   Button "Schaltfläche_256" at 1154,453 size 59x15; TextOff 'Text'
      on Click: SetTag("_DB_SDC_ERRORS.Error_nr", 830)
   Button "Schaltfläche_257" at 1154,469 size 59x15; TextOff 'Text'
      on Click: SetTag("_DB_SDC_ERRORS.Error_nr", 831)
   Button "Schaltfläche_258" at 1154,485 size 59x15; TextOff 'Text'
      on Click: SetTag("_DB_SDC_ERRORS.Error_nr", 832)
   Button "Schaltfläche_259" at 971,533 size 59x15; TextOff 'Text'
      on Click: SetTag("_DB_SDC_ERRORS.Error_nr", 901)
   Button "Schaltfläche_260" at 971,549 size 59x15; TextOff 'Text'
      on Click: SetTag("_DB_SDC_ERRORS.Error_nr", 902)
   Button "Schaltfläche_261" at 971,565 size 59x15; TextOff 'Text'
      on Click: SetTag("_DB_SDC_ERRORS.Error_nr", 903)
   Button "Schaltfläche_262" at 971,581 size 59x15; TextOff 'Text'
      on Click: SetTag("_DB_SDC_ERRORS.Error_nr", 904)
   Button "Schaltfläche_263" at 971,597 size 59x15; TextOff 'Text'
      on Click: SetTag("_DB_SDC_ERRORS.Error_nr", 905)
   Button "Schaltfläche_264" at 971,613 size 59x15; TextOff 'Text'
      on Click: SetTag("_DB_SDC_ERRORS.Error_nr", 906)
   Button "Schaltfläche_265" at 971,629 size 59x15; TextOff 'Text'
      on Click: SetTag("_DB_SDC_ERRORS.Error_nr", 907)
   Button "Schaltfläche_266" at 971,645 size 59x15; TextOff 'Text'
      on Click: SetTag("_DB_SDC_ERRORS.Error_nr", 908)
   Button "Schaltfläche_267" at 1033,533 size 59x15; TextOff 'Text'
      on Click: SetTag("_DB_SDC_ERRORS.Error_nr", 909)
   Button "Schaltfläche_268" at 1033,549 size 59x15; TextOff 'Text'
      on Click: SetTag("_DB_SDC_ERRORS.Error_nr", 910)
   Button "Schaltfläche_269" at 1033,565 size 59x15; TextOff 'Text'
      on Click: SetTag("_DB_SDC_ERRORS.Error_nr", 911)
   Button "Schaltfläche_270" at 1033,581 size 59x15; TextOff 'Text'
      on Click: SetTag("_DB_SDC_ERRORS.Error_nr", 912)
   Button "Schaltfläche_271" at 1033,597 size 59x15; TextOff 'Text'
      on Click: SetTag("_DB_SDC_ERRORS.Error_nr", 913)
   Button "Schaltfläche_272" at 1033,613 size 59x15; TextOff 'Text'
      on Click: SetTag("_DB_SDC_ERRORS.Error_nr", 914)
   Button "Schaltfläche_273" at 1033,629 size 59x15; TextOff 'Text'
      on Click: SetTag("_DB_SDC_ERRORS.Error_nr", 915)
   Button "Schaltfläche_274" at 1033,645 size 59x15; TextOff 'Text'
      on Click: SetTag("_DB_SDC_ERRORS.Error_nr", 916)
   Button "Schaltfläche_275" at 977,670 size 54x15; TextOff 'Text'
      on Click: SetTag("_DB_SDC_ERRORS.Error_nr", 917)
   Button "Schaltfläche_276" at 977,686 size 54x15; TextOff 'Text'
      on Click: SetTag("_DB_SDC_ERRORS.Error_nr", 918)
   Button "Schaltfläche_277" at 977,702 size 54x15; TextOff 'Text'
      on Click: SetTag("_DB_SDC_ERRORS.Error_nr", 919)
   Button "Schaltfläche_278" at 977,718 size 54x15; TextOff 'Text'
      on Click: SetTag("_DB_SDC_ERRORS.Error_nr", 920)
   Button "Schaltfläche_279" at 1032,669 size 54x15; TextOff 'Text'
      on Click: SetTag("_DB_SDC_ERRORS.Error_nr", 921)
   Button "Schaltfläche_280" at 1032,685 size 54x15; TextOff 'Text'
      on Click: SetTag("_DB_SDC_ERRORS.Error_nr", 922)
   Button "Schaltfläche_281" at 1032,701 size 54x15; TextOff 'Text'
      on Click: SetTag("_DB_SDC_ERRORS.Error_nr", 923)
   Button "Schaltfläche_282" at 1032,717 size 54x15; TextOff 'Text'
      on Click: SetTag("_DB_SDC_ERRORS.Error_nr", 924)

screen "724_ERROR_STAT_NOT_USED" 1280x800, template "Top_Header"
   on GenerateScreen: "SDC_ERROR_STAT"("SDC\DB_SDC_ERROR_STAT\_intern_Fault_Stat_Nr"); SetTag("SDC\_intern_Bildnummer", 724)
   IOField "EA-Feld_1" at 372,374 size 96x27; FormatPattern 999999999
      ProcessValue <- "SDC\DB_SDC_ERROR_STAT\DB_SDC_ERROR_STAT.F_STAT[XX1].EMS_TS_STAT_VAL.DRIVE_POS"
   TextField "Textfeld_1" at 353,331 size 170x27; Text 'Fahr-Pos [mm] / Drive Pos [mm] / Drive-Pos [mm]'
   IOField "EA-Feld_2" at 210,374 size 36x27; FormatPattern 999
      ProcessValue <- "SDC\DB_SDC_ERROR_STAT\DB_SDC_ERROR_STAT.F_STAT[XX1].EMS_TS_STAT_VAL.EMS_ID"
   TextField "Textfeld_2" at 195,331 size 80x27; Text 'EMS Nr'
   IOField "EA-Feld_3" at 676,374 size 36x27; FormatPattern 999
      ProcessValue <- "SDC\DB_SDC_ERROR_STAT\DB_SDC_ERROR_STAT.F_STAT[XX1].EMS_TS_STAT_VAL.ERROR"
   TextField "Textfeld_3" at 670,331 size 57x27; Text 'Error'
   IOField "EA-Feld_4" at 546,374 size 56x27; FormatPattern 99999
      ProcessValue <- "SDC\DB_SDC_ERROR_STAT\DB_SDC_ERROR_STAT.F_STAT[XX1].EMS_TS_STAT_VAL.HOIST_POS"
   TextField "Textfeld_4" at 506,331 size 169x27; Text 'Hub-Pos [mm] / Hoist Pos [mm]'
   IOField "EA-Feld_5" at 283,374 size 56x27; FormatPattern 99999
      ProcessValue <- "SDC\DB_SDC_ERROR_STAT\DB_SDC_ERROR_STAT.F_STAT[XX1].EMS_TS_STAT_VAL.SEK"
   TextField "Textfeld_5" at 273,331 size 83x27; Text 'Sektion / Section'
   TextField "Textfeld_6" at 988,331 size 155x27; Text 'date / time / Date and Time / Date / Time'
   Circle "Kreis_9" at 732,379 size 16x16
      Appearance <- "SDC\DB_SDC_ERROR_STAT\DB_SDC_ERROR_STAT.F_STAT[XX1].F"
   TextField "Textfeld_15" at 724,244 size 27x114; Text 'ER_BC_JUMP / F_BC_JUMP'
   Circle "Kreis_10" at 763,379 size 16x16
      Appearance <- "SDC\DB_SDC_ERROR_STAT\DB_SDC_ERROR_STAT.F_STAT[XX1].F"
   TextField "Textfeld_16" at 756,252 size 27x106; Text 'ER_NO_SEK / F_NO_SEK'
   Circle "Kreis_11" at 795,379 size 16x16
      Appearance <- "SDC\DB_SDC_ERROR_STAT\DB_SDC_ERROR_STAT.F_STAT[XX1].F"
   TextField "Textfeld_17" at 787,230 size 27x128; Text 'ER_COMMAND / F_COMMAND'
   Circle "Kreis_12" at 827,379 size 16x16
      Appearance <- "SDC\DB_SDC_ERROR_STAT\DB_SDC_ERROR_STAT.F_STAT[XX1].F"
   TextField "Textfeld_18" at 820,259 size 27x100; Text 'ER_BC_LIM / F_BC_LIM'
   Circle "Kreis_13" at 859,379 size 16x16
      Appearance <- "SDC\DB_SDC_ERROR_STAT\DB_SDC_ERROR_STAT.F_STAT[XX1].F"
   TextField "Textfeld_19" at 852,254 size 27x104; Text 'ER_EMS_ID / F_EMS_ID'
   Circle "Kreis_14" at 891,379 size 16x16
      Appearance <- "SDC\DB_SDC_ERROR_STAT\DB_SDC_ERROR_STAT.F_STAT[XX1].F"
   TextField "Textfeld_20" at 884,253 size 27x105; Text 'ER_SEK_NR / F_SEK_NR'
   Circle "Kreis_15" at 923,379 size 16x16
      Appearance <- "SDC\DB_SDC_ERROR_STAT\DB_SDC_ERROR_STAT.F_STAT[XX1].F"
   TextField "Textfeld_21" at 917,284 size 27x74; Text 'ER_LIFE / F_LIFE'
   Circle "Kreis_16" at 955,379 size 16x16
      Appearance <- "SDC\DB_SDC_ERROR_STAT\DB_SDC_ERROR_STAT.F_STAT[XX1].F"
   TextField "Textfeld_22" at 949,287 size 27x71; Text 'ER_BUS / F_BUS'
   TextField "Textfeld_23" at 425,169 size 127x27; Text 'pages / fehler entry / Error Entry'
   IOField "EA-Feld_8" at 151,374 size 36x27; FormatPattern 999
      ProcessValue <- "[0]"
   IOField "EA-Feld_9" at 372,414 size 96x27; FormatPattern 999999999
      ProcessValue <- "SDC\DB_SDC_ERROR_STAT\DB_SDC_ERROR_STAT.F_STAT[XX2].EMS_TS_STAT_VAL.DRIVE_POS"
   IOField "EA-Feld_10" at 210,414 size 36x27; FormatPattern 999
      ProcessValue <- "SDC\DB_SDC_ERROR_STAT\DB_SDC_ERROR_STAT.F_STAT[XX2].EMS_TS_STAT_VAL.EMS_ID"
   IOField "EA-Feld_11" at 676,414 size 36x27; FormatPattern 999
      ProcessValue <- "SDC\DB_SDC_ERROR_STAT\DB_SDC_ERROR_STAT.F_STAT[XX2].EMS_TS_STAT_VAL.ERROR"
   IOField "EA-Feld_12" at 546,414 size 56x27; FormatPattern 99999
      ProcessValue <- "SDC\DB_SDC_ERROR_STAT\DB_SDC_ERROR_STAT.F_STAT[XX2].EMS_TS_STAT_VAL.HOIST_POS"
   IOField "EA-Feld_13" at 283,414 size 56x27; FormatPattern 99999
      ProcessValue <- "SDC\DB_SDC_ERROR_STAT\DB_SDC_ERROR_STAT.F_STAT[XX2].EMS_TS_STAT_VAL.SEK"
   Circle "Kreis_17" at 732,419 size 16x16
      Appearance <- "SDC\DB_SDC_ERROR_STAT\DB_SDC_ERROR_STAT.F_STAT[XX2].F"
   Circle "Kreis_18" at 763,419 size 16x16
      Appearance <- "SDC\DB_SDC_ERROR_STAT\DB_SDC_ERROR_STAT.F_STAT[XX2].F"
   Circle "Kreis_19" at 795,419 size 16x16
      Appearance <- "SDC\DB_SDC_ERROR_STAT\DB_SDC_ERROR_STAT.F_STAT[XX2].F"
   Circle "Kreis_20" at 827,419 size 16x16
      Appearance <- "SDC\DB_SDC_ERROR_STAT\DB_SDC_ERROR_STAT.F_STAT[XX2].F"
   Circle "Kreis_21" at 859,419 size 16x16
      Appearance <- "SDC\DB_SDC_ERROR_STAT\DB_SDC_ERROR_STAT.F_STAT[XX2].F"
   Circle "Kreis_22" at 891,419 size 16x16
      Appearance <- "SDC\DB_SDC_ERROR_STAT\DB_SDC_ERROR_STAT.F_STAT[XX2].F"
   Circle "Kreis_23" at 923,419 size 16x16
      Appearance <- "SDC\DB_SDC_ERROR_STAT\DB_SDC_ERROR_STAT.F_STAT[XX2].F"
   Circle "Kreis_24" at 955,419 size 16x16
      Appearance <- "SDC\DB_SDC_ERROR_STAT\DB_SDC_ERROR_STAT.F_STAT[XX2].F"
   IOField "EA-Feld_15" at 151,414 size 36x27; FormatPattern 999
      ProcessValue <- "[1]"
   IOField "EA-Feld_16" at 372,454 size 96x27; FormatPattern 999999999
      ProcessValue <- "SDC\DB_SDC_ERROR_STAT\DB_SDC_ERROR_STAT.F_STAT[XX3].EMS_TS_STAT_VAL.DRIVE_POS"
   IOField "EA-Feld_17" at 210,454 size 36x27; FormatPattern 999
      ProcessValue <- "SDC\DB_SDC_ERROR_STAT\DB_SDC_ERROR_STAT.F_STAT[XX3].EMS_TS_STAT_VAL.EMS_ID"
   IOField "EA-Feld_18" at 676,454 size 36x27; FormatPattern 999
      ProcessValue <- "SDC\DB_SDC_ERROR_STAT\DB_SDC_ERROR_STAT.F_STAT[XX3].EMS_TS_STAT_VAL.ERROR"
   IOField "EA-Feld_19" at 546,454 size 56x27; FormatPattern 99999
      ProcessValue <- "SDC\DB_SDC_ERROR_STAT\DB_SDC_ERROR_STAT.F_STAT[XX3].EMS_TS_STAT_VAL.HOIST_POS"
   IOField "EA-Feld_20" at 283,454 size 56x27; FormatPattern 99999
      ProcessValue <- "SDC\DB_SDC_ERROR_STAT\DB_SDC_ERROR_STAT.F_STAT[XX3].EMS_TS_STAT_VAL.SEK"
   Circle "Kreis_25" at 732,459 size 16x16
      Appearance <- "SDC\DB_SDC_ERROR_STAT\DB_SDC_ERROR_STAT.F_STAT[XX3].F"
   Circle "Kreis_26" at 763,459 size 16x16
      Appearance <- "SDC\DB_SDC_ERROR_STAT\DB_SDC_ERROR_STAT.F_STAT[XX3].F"
   Circle "Kreis_27" at 795,459 size 16x16
      Appearance <- "SDC\DB_SDC_ERROR_STAT\DB_SDC_ERROR_STAT.F_STAT[XX3].F"
   Circle "Kreis_28" at 827,459 size 16x16
      Appearance <- "SDC\DB_SDC_ERROR_STAT\DB_SDC_ERROR_STAT.F_STAT[XX3].F"
   Circle "Kreis_29" at 859,459 size 16x16
      Appearance <- "SDC\DB_SDC_ERROR_STAT\DB_SDC_ERROR_STAT.F_STAT[XX3].F"
   Circle "Kreis_30" at 891,459 size 16x16
      Appearance <- "SDC\DB_SDC_ERROR_STAT\DB_SDC_ERROR_STAT.F_STAT[XX3].F"
   Circle "Kreis_31" at 923,459 size 16x16
      Appearance <- "SDC\DB_SDC_ERROR_STAT\DB_SDC_ERROR_STAT.F_STAT[XX3].F"
   Circle "Kreis_32" at 955,459 size 16x16
      Appearance <- "SDC\DB_SDC_ERROR_STAT\DB_SDC_ERROR_STAT.F_STAT[XX3].F"
   IOField "EA-Feld_22" at 151,454 size 36x27; FormatPattern 999
      ProcessValue <- "[2]"
   IOField "EA-Feld_23" at 372,494 size 96x27; FormatPattern 999999999
      ProcessValue <- "SDC\DB_SDC_ERROR_STAT\DB_SDC_ERROR_STAT.F_STAT[XX4].EMS_TS_STAT_VAL.DRIVE_POS"
   IOField "EA-Feld_24" at 210,494 size 36x27; FormatPattern 999
      ProcessValue <- "SDC\DB_SDC_ERROR_STAT\DB_SDC_ERROR_STAT.F_STAT[XX4].EMS_TS_STAT_VAL.EMS_ID"
   IOField "EA-Feld_25" at 676,494 size 36x27; FormatPattern 999
      ProcessValue <- "SDC\DB_SDC_ERROR_STAT\DB_SDC_ERROR_STAT.F_STAT[XX4].EMS_TS_STAT_VAL.ERROR"
   IOField "EA-Feld_26" at 546,494 size 56x27; FormatPattern 99999
      ProcessValue <- "SDC\DB_SDC_ERROR_STAT\DB_SDC_ERROR_STAT.F_STAT[XX4].EMS_TS_STAT_VAL.HOIST_POS"
   IOField "EA-Feld_27" at 283,494 size 56x27; FormatPattern 99999
      ProcessValue <- "SDC\DB_SDC_ERROR_STAT\DB_SDC_ERROR_STAT.F_STAT[XX4].EMS_TS_STAT_VAL.SEK"
   Circle "Kreis_33" at 732,499 size 16x16
      Appearance <- "SDC\DB_SDC_ERROR_STAT\DB_SDC_ERROR_STAT.F_STAT[XX4].F"
   Circle "Kreis_34" at 763,499 size 16x16
      Appearance <- "SDC\DB_SDC_ERROR_STAT\DB_SDC_ERROR_STAT.F_STAT[XX4].F"
   Circle "Kreis_35" at 795,499 size 16x16
      Appearance <- "SDC\DB_SDC_ERROR_STAT\DB_SDC_ERROR_STAT.F_STAT[XX4].F"
   Circle "Kreis_36" at 827,499 size 16x16
      Appearance <- "SDC\DB_SDC_ERROR_STAT\DB_SDC_ERROR_STAT.F_STAT[XX4].F"
   Circle "Kreis_37" at 859,499 size 16x16
      Appearance <- "SDC\DB_SDC_ERROR_STAT\DB_SDC_ERROR_STAT.F_STAT[XX4].F"
   Circle "Kreis_38" at 891,499 size 16x16
      Appearance <- "SDC\DB_SDC_ERROR_STAT\DB_SDC_ERROR_STAT.F_STAT[XX4].F"
   Circle "Kreis_39" at 923,499 size 16x16
      Appearance <- "SDC\DB_SDC_ERROR_STAT\DB_SDC_ERROR_STAT.F_STAT[XX4].F"
   Circle "Kreis_40" at 955,499 size 16x16
      Appearance <- "SDC\DB_SDC_ERROR_STAT\DB_SDC_ERROR_STAT.F_STAT[XX4].F"
   IOField "EA-Feld_29" at 151,494 size 36x27; FormatPattern 999
      ProcessValue <- "[3]"
   IOField "EA-Feld_30" at 372,534 size 96x27; FormatPattern 999999999
      ProcessValue <- "SDC\DB_SDC_ERROR_STAT\DB_SDC_ERROR_STAT.F_STAT[XX5].EMS_TS_STAT_VAL.DRIVE_POS"
   IOField "EA-Feld_31" at 210,534 size 36x27; FormatPattern 999
      ProcessValue <- "SDC\DB_SDC_ERROR_STAT\DB_SDC_ERROR_STAT.F_STAT[XX5].EMS_TS_STAT_VAL.EMS_ID"
   IOField "EA-Feld_32" at 676,534 size 36x27; FormatPattern 999
      ProcessValue <- "SDC\DB_SDC_ERROR_STAT\DB_SDC_ERROR_STAT.F_STAT[XX5].EMS_TS_STAT_VAL.ERROR"
   IOField "EA-Feld_33" at 546,534 size 56x27; FormatPattern 99999
      ProcessValue <- "SDC\DB_SDC_ERROR_STAT\DB_SDC_ERROR_STAT.F_STAT[XX5].EMS_TS_STAT_VAL.HOIST_POS"
   IOField "EA-Feld_34" at 283,534 size 56x27; FormatPattern 99999
      ProcessValue <- "SDC\DB_SDC_ERROR_STAT\DB_SDC_ERROR_STAT.F_STAT[XX5].EMS_TS_STAT_VAL.SEK"
   Circle "Kreis_41" at 732,539 size 16x16
      Appearance <- "SDC\DB_SDC_ERROR_STAT\DB_SDC_ERROR_STAT.F_STAT[XX5].F"
   Circle "Kreis_42" at 763,539 size 16x16
      Appearance <- "SDC\DB_SDC_ERROR_STAT\DB_SDC_ERROR_STAT.F_STAT[XX5].F"
   Circle "Kreis_43" at 795,539 size 16x16
      Appearance <- "SDC\DB_SDC_ERROR_STAT\DB_SDC_ERROR_STAT.F_STAT[XX5].F"
   Circle "Kreis_44" at 827,539 size 16x16
      Appearance <- "SDC\DB_SDC_ERROR_STAT\DB_SDC_ERROR_STAT.F_STAT[XX5].F"
   Circle "Kreis_45" at 859,539 size 16x16
      Appearance <- "SDC\DB_SDC_ERROR_STAT\DB_SDC_ERROR_STAT.F_STAT[XX5].F"
   Circle "Kreis_46" at 891,539 size 16x16
      Appearance <- "SDC\DB_SDC_ERROR_STAT\DB_SDC_ERROR_STAT.F_STAT[XX5].F"
   Circle "Kreis_47" at 923,539 size 16x16
      Appearance <- "SDC\DB_SDC_ERROR_STAT\DB_SDC_ERROR_STAT.F_STAT[XX5].F"
   Circle "Kreis_48" at 955,539 size 16x16
      Appearance <- "SDC\DB_SDC_ERROR_STAT\DB_SDC_ERROR_STAT.F_STAT[XX5].F"
   IOField "EA-Feld_36" at 151,534 size 36x27; FormatPattern 999
      ProcessValue <- "[4]"
   IOField "EA-Feld_37" at 372,574 size 96x27; FormatPattern 999999999
      ProcessValue <- "SDC\DB_SDC_ERROR_STAT\DB_SDC_ERROR_STAT.F_STAT[XX6].EMS_TS_STAT_VAL.DRIVE_POS"
   IOField "EA-Feld_38" at 210,574 size 36x27; FormatPattern 999
      ProcessValue <- "SDC\DB_SDC_ERROR_STAT\DB_SDC_ERROR_STAT.F_STAT[XX6].EMS_TS_STAT_VAL.EMS_ID"
   IOField "EA-Feld_39" at 676,574 size 36x27; FormatPattern 999
      ProcessValue <- "SDC\DB_SDC_ERROR_STAT\DB_SDC_ERROR_STAT.F_STAT[XX6].EMS_TS_STAT_VAL.ERROR"
   IOField "EA-Feld_40" at 546,574 size 56x27; FormatPattern 99999
      ProcessValue <- "SDC\DB_SDC_ERROR_STAT\DB_SDC_ERROR_STAT.F_STAT[XX6].EMS_TS_STAT_VAL.HOIST_POS"
   IOField "EA-Feld_41" at 283,574 size 56x27; FormatPattern 99999
      ProcessValue <- "SDC\DB_SDC_ERROR_STAT\DB_SDC_ERROR_STAT.F_STAT[XX6].EMS_TS_STAT_VAL.SEK"
   Circle "Kreis_49" at 732,579 size 16x16
      Appearance <- "SDC\DB_SDC_ERROR_STAT\DB_SDC_ERROR_STAT.F_STAT[XX6].F"
   Circle "Kreis_50" at 763,579 size 16x16
      Appearance <- "SDC\DB_SDC_ERROR_STAT\DB_SDC_ERROR_STAT.F_STAT[XX6].F"
   Circle "Kreis_51" at 795,579 size 16x16
      Appearance <- "SDC\DB_SDC_ERROR_STAT\DB_SDC_ERROR_STAT.F_STAT[XX6].F"
   Circle "Kreis_52" at 827,579 size 16x16
      Appearance <- "SDC\DB_SDC_ERROR_STAT\DB_SDC_ERROR_STAT.F_STAT[XX6].F"
   Circle "Kreis_53" at 859,579 size 16x16
      Appearance <- "SDC\DB_SDC_ERROR_STAT\DB_SDC_ERROR_STAT.F_STAT[XX6].F"
   Circle "Kreis_54" at 891,579 size 16x16
      Appearance <- "SDC\DB_SDC_ERROR_STAT\DB_SDC_ERROR_STAT.F_STAT[XX6].F"
   Circle "Kreis_55" at 923,579 size 16x16
      Appearance <- "SDC\DB_SDC_ERROR_STAT\DB_SDC_ERROR_STAT.F_STAT[XX6].F"
   Circle "Kreis_56" at 955,579 size 16x16
      Appearance <- "SDC\DB_SDC_ERROR_STAT\DB_SDC_ERROR_STAT.F_STAT[XX6].F"
   IOField "EA-Feld_43" at 151,574 size 36x27; FormatPattern 999
      ProcessValue <- "[5]"
   IOField "EA-Feld_44" at 372,614 size 96x27; FormatPattern 999999999
      ProcessValue <- "SDC\DB_SDC_ERROR_STAT\DB_SDC_ERROR_STAT.F_STAT[XX7].EMS_TS_STAT_VAL.DRIVE_POS"
   IOField "EA-Feld_45" at 210,614 size 36x27; FormatPattern 999
      ProcessValue <- "SDC\DB_SDC_ERROR_STAT\DB_SDC_ERROR_STAT.F_STAT[XX7].EMS_TS_STAT_VAL.EMS_ID"
   IOField "EA-Feld_46" at 676,614 size 36x27; FormatPattern 999
      ProcessValue <- "SDC\DB_SDC_ERROR_STAT\DB_SDC_ERROR_STAT.F_STAT[XX7].EMS_TS_STAT_VAL.ERROR"
   IOField "EA-Feld_47" at 546,614 size 56x27; FormatPattern 99999
      ProcessValue <- "SDC\DB_SDC_ERROR_STAT\DB_SDC_ERROR_STAT.F_STAT[XX7].EMS_TS_STAT_VAL.HOIST_POS"
   IOField "EA-Feld_48" at 283,614 size 56x27; FormatPattern 99999
      ProcessValue <- "SDC\DB_SDC_ERROR_STAT\DB_SDC_ERROR_STAT.F_STAT[XX7].EMS_TS_STAT_VAL.SEK"
   Circle "Kreis_57" at 732,619 size 16x16
      Appearance <- "SDC\DB_SDC_ERROR_STAT\DB_SDC_ERROR_STAT.F_STAT[XX7].F"
   Circle "Kreis_58" at 763,619 size 16x16
      Appearance <- "SDC\DB_SDC_ERROR_STAT\DB_SDC_ERROR_STAT.F_STAT[XX7].F"
   Circle "Kreis_59" at 795,619 size 16x16
      Appearance <- "SDC\DB_SDC_ERROR_STAT\DB_SDC_ERROR_STAT.F_STAT[XX7].F"
   Circle "Kreis_60" at 827,619 size 16x16
      Appearance <- "SDC\DB_SDC_ERROR_STAT\DB_SDC_ERROR_STAT.F_STAT[XX7].F"
   Circle "Kreis_61" at 859,619 size 16x16
      Appearance <- "SDC\DB_SDC_ERROR_STAT\DB_SDC_ERROR_STAT.F_STAT[XX7].F"
   Circle "Kreis_62" at 891,619 size 16x16
      Appearance <- "SDC\DB_SDC_ERROR_STAT\DB_SDC_ERROR_STAT.F_STAT[XX7].F"
   Circle "Kreis_63" at 923,619 size 16x16
      Appearance <- "SDC\DB_SDC_ERROR_STAT\DB_SDC_ERROR_STAT.F_STAT[XX7].F"
   Circle "Kreis_64" at 955,619 size 16x16
      Appearance <- "SDC\DB_SDC_ERROR_STAT\DB_SDC_ERROR_STAT.F_STAT[XX7].F"
   IOField "EA-Feld_50" at 151,614 size 36x27; FormatPattern 999
      ProcessValue <- "[6]"
   IOField "EA-Feld_51" at 372,654 size 96x27; FormatPattern 999999999
      ProcessValue <- "SDC\DB_SDC_ERROR_STAT\DB_SDC_ERROR_STAT.F_STAT[XX8].EMS_TS_STAT_VAL.DRIVE_POS"
   IOField "EA-Feld_52" at 210,654 size 36x27; FormatPattern 999
      ProcessValue <- "SDC\DB_SDC_ERROR_STAT\DB_SDC_ERROR_STAT.F_STAT[XX8].EMS_TS_STAT_VAL.EMS_ID"
   IOField "EA-Feld_53" at 676,654 size 36x27; FormatPattern 999
      ProcessValue <- "SDC\DB_SDC_ERROR_STAT\DB_SDC_ERROR_STAT.F_STAT[XX8].EMS_TS_STAT_VAL.ERROR"
   IOField "EA-Feld_54" at 546,654 size 56x27; FormatPattern 99999
      ProcessValue <- "SDC\DB_SDC_ERROR_STAT\DB_SDC_ERROR_STAT.F_STAT[XX8].EMS_TS_STAT_VAL.HOIST_POS"
   IOField "EA-Feld_55" at 283,654 size 56x27; FormatPattern 99999
      ProcessValue <- "SDC\DB_SDC_ERROR_STAT\DB_SDC_ERROR_STAT.F_STAT[XX8].EMS_TS_STAT_VAL.SEK"
   Circle "Kreis_65" at 732,659 size 16x16
      Appearance <- "SDC\DB_SDC_ERROR_STAT\DB_SDC_ERROR_STAT.F_STAT[XX8].F"
   Circle "Kreis_66" at 763,659 size 16x16
      Appearance <- "SDC\DB_SDC_ERROR_STAT\DB_SDC_ERROR_STAT.F_STAT[XX8].F"
   Circle "Kreis_67" at 795,659 size 16x16
      Appearance <- "SDC\DB_SDC_ERROR_STAT\DB_SDC_ERROR_STAT.F_STAT[XX8].F"
   Circle "Kreis_68" at 827,659 size 16x16
      Appearance <- "SDC\DB_SDC_ERROR_STAT\DB_SDC_ERROR_STAT.F_STAT[XX8].F"
   Circle "Kreis_69" at 859,659 size 16x16
      Appearance <- "SDC\DB_SDC_ERROR_STAT\DB_SDC_ERROR_STAT.F_STAT[XX8].F"
   Circle "Kreis_70" at 891,659 size 16x16
      Appearance <- "SDC\DB_SDC_ERROR_STAT\DB_SDC_ERROR_STAT.F_STAT[XX8].F"
   Circle "Kreis_71" at 923,659 size 16x16
      Appearance <- "SDC\DB_SDC_ERROR_STAT\DB_SDC_ERROR_STAT.F_STAT[XX8].F"
   Circle "Kreis_72" at 955,659 size 16x16
      Appearance <- "SDC\DB_SDC_ERROR_STAT\DB_SDC_ERROR_STAT.F_STAT[XX8].F"
   IOField "EA-Feld_57" at 151,654 size 36x27; FormatPattern 999
      ProcessValue <- "[7]"
   IOField "EA-Feld_58" at 372,694 size 96x27; FormatPattern 999999999
      ProcessValue <- "SDC\DB_SDC_ERROR_STAT\DB_SDC_ERROR_STAT.F_STAT[XX9].EMS_TS_STAT_VAL.DRIVE_POS"
   IOField "EA-Feld_59" at 210,694 size 36x27; FormatPattern 999
      ProcessValue <- "SDC\DB_SDC_ERROR_STAT\DB_SDC_ERROR_STAT.F_STAT[XX9].EMS_TS_STAT_VAL.EMS_ID"
   IOField "EA-Feld_60" at 676,694 size 36x27; FormatPattern 999
      ProcessValue <- "SDC\DB_SDC_ERROR_STAT\DB_SDC_ERROR_STAT.F_STAT[XX9].EMS_TS_STAT_VAL.ERROR"
   IOField "EA-Feld_61" at 546,694 size 56x27; FormatPattern 99999
      ProcessValue <- "SDC\DB_SDC_ERROR_STAT\DB_SDC_ERROR_STAT.F_STAT[XX9].EMS_TS_STAT_VAL.HOIST_POS"
   IOField "EA-Feld_62" at 283,694 size 56x27; FormatPattern 99999
      ProcessValue <- "SDC\DB_SDC_ERROR_STAT\DB_SDC_ERROR_STAT.F_STAT[XX9].EMS_TS_STAT_VAL.SEK"
   Circle "Kreis_73" at 732,699 size 16x16
      Appearance <- "SDC\DB_SDC_ERROR_STAT\DB_SDC_ERROR_STAT.F_STAT[XX9].F"
   Circle "Kreis_74" at 763,699 size 16x16
      Appearance <- "SDC\DB_SDC_ERROR_STAT\DB_SDC_ERROR_STAT.F_STAT[XX9].F"
   Circle "Kreis_75" at 795,699 size 16x16
      Appearance <- "SDC\DB_SDC_ERROR_STAT\DB_SDC_ERROR_STAT.F_STAT[XX9].F"
   Circle "Kreis_76" at 827,699 size 16x16
      Appearance <- "SDC\DB_SDC_ERROR_STAT\DB_SDC_ERROR_STAT.F_STAT[XX9].F"
   Circle "Kreis_77" at 859,699 size 16x16
      Appearance <- "SDC\DB_SDC_ERROR_STAT\DB_SDC_ERROR_STAT.F_STAT[XX9].F"
   Circle "Kreis_78" at 891,699 size 16x16
      Appearance <- "SDC\DB_SDC_ERROR_STAT\DB_SDC_ERROR_STAT.F_STAT[XX9].F"
   Circle "Kreis_79" at 923,699 size 16x16
      Appearance <- "SDC\DB_SDC_ERROR_STAT\DB_SDC_ERROR_STAT.F_STAT[XX9].F"
   Circle "Kreis_80" at 955,699 size 16x16
      Appearance <- "SDC\DB_SDC_ERROR_STAT\DB_SDC_ERROR_STAT.F_STAT[XX9].F"
   IOField "EA-Feld_64" at 151,694 size 36x27; FormatPattern 999
      ProcessValue <- "[8]"
   IOField "EA-Feld_65" at 372,734 size 96x27; FormatPattern 999999999
      ProcessValue <- "SDC\DB_SDC_ERROR_STAT\DB_SDC_ERROR_STAT.F_STAT[X10].EMS_TS_STAT_VAL.DRIVE_POS"
   IOField "EA-Feld_66" at 210,734 size 36x27; FormatPattern 999
      ProcessValue <- "SDC\DB_SDC_ERROR_STAT\DB_SDC_ERROR_STAT.F_STAT[X10].EMS_TS_STAT_VAL.EMS_ID"
   IOField "EA-Feld_67" at 676,734 size 36x27; FormatPattern 999
      ProcessValue <- "SDC\DB_SDC_ERROR_STAT\DB_SDC_ERROR_STAT.F_STAT[X10].EMS_TS_STAT_VAL.ERROR"
   IOField "EA-Feld_68" at 546,734 size 56x27; FormatPattern 99999
      ProcessValue <- "SDC\DB_SDC_ERROR_STAT\DB_SDC_ERROR_STAT.F_STAT[X10].EMS_TS_STAT_VAL.HOIST_POS"
   IOField "EA-Feld_69" at 283,734 size 56x27; FormatPattern 99999
      ProcessValue <- "SDC\DB_SDC_ERROR_STAT\DB_SDC_ERROR_STAT.F_STAT[X10].EMS_TS_STAT_VAL.SEK"
   Circle "Kreis_81" at 732,739 size 16x16
      Appearance <- "SDC\DB_SDC_ERROR_STAT\DB_SDC_ERROR_STAT.F_STAT[X10].F"
   Circle "Kreis_82" at 763,739 size 16x16
      Appearance <- "SDC\DB_SDC_ERROR_STAT\DB_SDC_ERROR_STAT.F_STAT[X10].F"
   Circle "Kreis_83" at 795,739 size 16x16
      Appearance <- "SDC\DB_SDC_ERROR_STAT\DB_SDC_ERROR_STAT.F_STAT[X10].F"
   Circle "Kreis_84" at 827,739 size 16x16
      Appearance <- "SDC\DB_SDC_ERROR_STAT\DB_SDC_ERROR_STAT.F_STAT[X10].F"
   Circle "Kreis_85" at 859,739 size 16x16
      Appearance <- "SDC\DB_SDC_ERROR_STAT\DB_SDC_ERROR_STAT.F_STAT[X10].F"
   Circle "Kreis_86" at 891,739 size 16x16
      Appearance <- "SDC\DB_SDC_ERROR_STAT\DB_SDC_ERROR_STAT.F_STAT[X10].F"
   Circle "Kreis_87" at 923,739 size 16x16
      Appearance <- "SDC\DB_SDC_ERROR_STAT\DB_SDC_ERROR_STAT.F_STAT[X10].F"
   Circle "Kreis_88" at 955,739 size 16x16
      Appearance <- "SDC\DB_SDC_ERROR_STAT\DB_SDC_ERROR_STAT.F_STAT[X10].F"
   IOField "EA-Feld_71" at 151,734 size 36x27; FormatPattern 999
      ProcessValue <- "[9]"
   Button "Schaltfläche_1" at 374,166 size 40x32; TextOff '+'
      on Click: function_dd21b452("SDC\DB_SDC_ERROR_STAT\_intern_Fault_Stat_Nr", 10); "SDC_ERROR_STAT"("SDC\DB_SDC_ERROR_STAT\_intern_Fault_Stat_Nr")
   Button "Schaltfläche_3" at 277,166 size 39x32; TextOff '-'
      on Click: function_b9b71300("SDC\DB_SDC_ERROR_STAT\_intern_Fault_Stat_Nr", 10); "SDC_ERROR_STAT"("SDC\DB_SDC_ERROR_STAT\_intern_Fault_Stat_Nr")
   IOField "EA-Feld_7" at 317,166 size 56x32; FormatPattern 9999
      on OnFinishInput: "SDC_ERROR_STAT"("SDC\DB_SDC_ERROR_STAT\_intern_Fault_Stat_Nr")
      ProcessValue <- "SDC\DB_SDC_ERROR_STAT\_intern_Fault_Stat_Nr"
   TextField "Textfeld_24" at 657,169 size 234x27; Text 'max. count / maximum fault entrys / Max. Error Messages'
   IOField "EA-Feld_72" at 589,166 size 56x32; FormatPattern 9999
      on OnFinishInput: "SDC_ERROR_STAT"("SDC\DB_SDC_ERROR_STAT\_intern_Fault_Stat_Nr")
      Appearance <- "SDC\_EDIT"
      ObjectEnable <- "SDC\_EDIT"
      ProcessValue <- "DB_SDC_ERRORS_STAT_HEADER.MAX_NR_FAULT_STAT"
   Button "Schaltfläche_38" at 3,712 size 127x84; TextOff 'EDIT'
      on Click: SetTag("SDC\_EDIT", 1); InvertBit("SDC\_EDIT_BIT")
      Appearance <- "SDC\_EDIT"
   Button "Schaltfläche_42" at 3,712 size 127x84; TextOff 'EDIT'
      on Click: SetTag("SDC\_EDIT", 0); InvertBit("SDC\_EDIT_BIT")
      Visibility <- "SDC\_EDIT"
      Appearance <- "SDC\_EDIT"
   Button "Schaltfläche_2" at 866,169 size 299x31; TextOff 'delete archive / EDIT / Delete Archieve'
      on Click: SetBit("DB_SDC_ERRORS_STAT_HEADER.RESET_ARCH")
      on Release: ResetBit("DB_SDC_ERRORS_STAT_HEADER.RESET_ARCH")
      Visibility <- "SDC\_EDIT"
   IOField "EA-Feld_6" at 988,374 size 212x27
      ProcessValue <- "SDC\DB_SDC_ERROR_STAT\DB_SDC_ERROR_STAT.F_STAT[XX1].F_DATE"
   IOField "EA-Feld_14" at 988,414 size 212x27
      ProcessValue <- "SDC\DB_SDC_ERROR_STAT\DB_SDC_ERROR_STAT.F_STAT[XX2].F_DATE"
   IOField "EA-Feld_21" at 988,454 size 212x27
      ProcessValue <- "SDC\DB_SDC_ERROR_STAT\DB_SDC_ERROR_STAT.F_STAT[XX3].F_DATE"
   IOField "EA-Feld_28" at 988,494 size 212x27
      ProcessValue <- "SDC\DB_SDC_ERROR_STAT\DB_SDC_ERROR_STAT.F_STAT[XX4].F_DATE"
   IOField "EA-Feld_35" at 988,534 size 212x27
      ProcessValue <- "SDC\DB_SDC_ERROR_STAT\DB_SDC_ERROR_STAT.F_STAT[XX5].F_DATE"
   IOField "EA-Feld_42" at 988,574 size 212x27
      ProcessValue <- "SDC\DB_SDC_ERROR_STAT\DB_SDC_ERROR_STAT.F_STAT[XX6].F_DATE"
   IOField "EA-Feld_49" at 988,614 size 212x27
      ProcessValue <- "SDC\DB_SDC_ERROR_STAT\DB_SDC_ERROR_STAT.F_STAT[XX7].F_DATE"
   IOField "EA-Feld_56" at 988,654 size 212x27
      ProcessValue <- "SDC\DB_SDC_ERROR_STAT\DB_SDC_ERROR_STAT.F_STAT[XX8].F_DATE"
   IOField "EA-Feld_63" at 988,694 size 212x27
      ProcessValue <- "SDC\DB_SDC_ERROR_STAT\DB_SDC_ERROR_STAT.F_STAT[XX9].F_DATE"
   IOField "EA-Feld_70" at 988,734 size 212x27
      ProcessValue <- "SDC\DB_SDC_ERROR_STAT\DB_SDC_ERROR_STAT.F_STAT[X10].F_DATE"

screen "728_CARRIER_VFD_STATUS" 1280x800, template "Top_Header"
   on GenerateScreen: "SDC_EMS_STATUS"('SDC\DB_SDC_EMS\_Intern_EMS_Nr'); "SDC_TS_REFERENCE"("SDC\DB_SDC_EMS\EMS[XXX].TS_STAT.VAL.SEK"); SetTag("SDC\DB_SDC_EMS\HMI[XX].BILD_Nr", 728); "SDC_EMS_TA_STATUS"("HMI_EMS_Nr"); SetTag("SDC\_intern_Bildnummer", 728)
   on ClearScreen: SetTag("SDC\DB_SDC_EMS\HMI[XX].BILD_Nr", 0)
   IOField "EA-Feld_4" at 261,138 size 56x32; FormatPattern 9999
      on OnFinishInput: "SDC_EMS_STATUS"("HMI_EMS_Nr"); "SDC_EMS_TA_STATUS"("HMI_EMS_Nr")
      ProcessValue <- "HMI_EMS_Nr"
   TextField "Textfeld_3" at 369,141 size 100x25; Text 'EMS-No. / EMS-Number / Carrier-No.'
   Button "Schaltfläche_1" at 318,138 size 40x32; TextOff '+'
      on Click: function_dd21b452("HMI_EMS_Nr", 1); "SDC_EMS_STATUS"("HMI_EMS_Nr"); "SDC_EMS_TA_STATUS"("HMI_EMS_Nr")
   Button "Schaltfläche_3" at 221,138 size 39x32; TextOff '-'
      on Click: function_b9b71300("HMI_EMS_Nr", 1); "SDC_EMS_STATUS"("HMI_EMS_Nr"); "SDC_EMS_TA_STATUS"("HMI_EMS_Nr")
   SymbolicIOField "Symbolisches EA-Feld_2" at 205,698 size 901x26; TextOn '1'; TextOff '0'; TextList "G120D_Faults_Warnings"
      ProcessValue <- "DB_SDC_EMS_TA.EMS[XX].TA1.FAULT"
   SymbolicIOField "Symbolisches EA-Feld_1" at 205,743 size 901x26; TextOn '1'; TextOff '0'; TextList "G120D_Faults_Warnings"
      ProcessValue <- "DB_SDC_EMS_TA.EMS[XX].TA1.ALARM"
   TextField "Textfeld_1" at 558,118 size 243x27; Text 'section counter / min Barcode mm / Carrier Drive Status'
   TextField "Text field_1" at 219,197 size 274x25; Text 'G120 DRIVE STW1 CONTROL'
   TextField "Text field_2" at 819,203 size 259x25; Text 'G120 DRIVE ZSW1 STATUS'
   TextField "Textfeld_2" at 241,241 size 100x25; Text 'EMS-No. / EMS-Number / ON'
   TextField "Textfeld_4" at 241,266 size 100x25; Text 'EMS-No. / EMS-Number / AUS2_INH'
   TextField "Textfeld_5" at 241,291 size 100x25; Text 'EMS-No. / EMS-Number / AUS3_STOP'
   TextField "Textfeld_6" at 241,316 size 100x25; Text 'EMS-No. / EMS-Number / ENABLE'
   TextField "Textfeld_7" at 241,341 size 113x25; Text 'EMS-No. / EMS-Number / ENABLE RAMP'
   TextField "Textfeld_8" at 241,366 size 104x25; Text 'EMS-No. / EMS-Number / START RAMP'
   TextField "Textfeld_9" at 241,391 size 100x25; Text 'EMS-No. / EMS-Number / SET POINT'
   TextField "Textfeld_10" at 241,416 size 100x25; Text 'EMS-No. / EMS-Number / RESET'
   TextField "Textfeld_11" at 241,441 size 100x25; Text 'EMS-No. / EMS-Number / JOG RIGHT'
   TextField "Textfeld_12" at 241,466 size 100x25; Text 'EMS-No. / EMS-Number / JOG LEFT'
   TextField "Textfeld_13" at 241,491 size 110x25; Text 'EMS-No. / EMS-Number / CONTROL PLC'
   TextField "Textfeld_14" at 241,516 size 100x25; Text 'EMS-No. / EMS-Number / REVERSE'
   TextField "Textfeld_15" at 241,541 size 130x25; Text 'EMS-No. / EMS-Number / BRAKE RELEASE'
   TextField "Textfeld_16" at 241,566 size 100x25; Text 'EMS-No. / EMS-Number / DDS'
   TextField "Textfeld_17" at 241,591 size 100x25; Text 'EMS-No. / EMS-Number / DO0'
   TextField "Textfeld_18" at 241,616 size 100x25; Text 'EMS-No. / EMS-Number / DO1'
   TextField "Textfeld_19" at 834,248 size 100x25; Text 'EMS-No. / EMS-Number / READY RUN'
   TextField "Textfeld_20" at 834,273 size 100x25; Text 'EMS-No. / EMS-Number / READY ON'
   TextField "Textfeld_21" at 834,298 size 100x25; Text 'EMS-No. / EMS-Number / ENABLE'
   TextField "Textfeld_22" at 834,323 size 100x25; Text 'EMS-No. / EMS-Number / FAULT'
   TextField "Textfeld_23" at 834,348 size 100x25; Text 'EMS-No. / EMS-Number / OFF 2'
   TextField "Textfeld_24" at 834,373 size 100x25; Text 'EMS-No. / EMS-Number / OFF 3'
   TextField "Textfeld_25" at 834,398 size 100x25; Text 'EMS-No. / EMS-Number / LOCK OUT'
   TextField "Textfeld_26" at 834,423 size 100x25; Text 'EMS-No. / EMS-Number / WARN'
   TextField "Textfeld_27" at 834,448 size 120x25; Text 'EMS-No. / EMS-Number / NO DEVIATION'
   TextField "Textfeld_28" at 834,473 size 110x25; Text 'EMS-No. / EMS-Number / CONTROL PLC'
   TextField "Textfeld_29" at 834,498 size 100x25; Text 'EMS-No. / EMS-Number / F MAX'
   TextField "Textfeld_30" at 834,523 size 127x25; Text 'EMS-No. / EMS-Number / LIMIT REACHED'
   TextField "Textfeld_31" at 834,548 size 103x25; Text 'EMS-No. / EMS-Number / BRAKE OPEN'
   TextField "Textfeld_32" at 834,573 size 117x25; Text 'EMS-No. / EMS-Number / NO OVERTEMP'
   TextField "Textfeld_33" at 834,598 size 100x25; Text 'EMS-No. / EMS-Number / CW_CCW'
   TextField "Textfeld_34" at 834,621 size 100x25; Text 'EMS-No. / EMS-Number / OVERLOAD'
   Circle "Kreis_15" at 220,246 size 15x15
      Appearance <- "HMI_Status_G120D_Control"
   Circle "Kreis_1" at 220,271 size 15x15
      Appearance <- "HMI_Status_G120D_Control"
   Circle "Kreis_2" at 220,296 size 15x15
      Appearance <- "HMI_Status_G120D_Control"
   Circle "Kreis_3" at 220,321 size 15x15
      Appearance <- "HMI_Status_G120D_Control"
   Circle "Kreis_4" at 220,346 size 15x15
      Appearance <- "HMI_Status_G120D_Control"
   Circle "Kreis_5" at 220,371 size 15x15
      Appearance <- "HMI_Status_G120D_Control"
   Circle "Kreis_6" at 220,396 size 15x15
      Appearance <- "HMI_Status_G120D_Control"
   Circle "Kreis_7" at 220,421 size 15x15
      Appearance <- "HMI_Status_G120D_Control"
   Circle "Kreis_8" at 220,446 size 15x15
      Appearance <- "HMI_Status_G120D_Control"
   Circle "Kreis_9" at 220,471 size 15x15
      Appearance <- "HMI_Status_G120D_Control"
   Circle "Kreis_10" at 220,496 size 15x15
      Appearance <- "HMI_Status_G120D_Control"
   Circle "Kreis_11" at 220,521 size 15x15
      Appearance <- "HMI_Status_G120D_Control"
   Circle "Kreis_12" at 220,546 size 15x15
      Appearance <- "HMI_Status_G120D_Control"
   Circle "Kreis_13" at 220,571 size 15x15
      Appearance <- "HMI_Status_G120D_Control"
   Circle "Kreis_14" at 220,596 size 15x15
      Appearance <- "HMI_Status_G120D_Control"
   Circle "Kreis_16" at 220,621 size 15x15
      Appearance <- "HMI_Status_G120D_Control"
   Circle "Kreis_17" at 813,253 size 15x15
      Appearance <- "HMI_Status_G120D_Status"
   Circle "Kreis_18" at 813,278 size 15x15
      Appearance <- "HMI_Status_G120D_Status"
   Circle "Kreis_19" at 813,303 size 15x15
      Appearance <- "HMI_Status_G120D_Status"
   Circle "Kreis_20" at 813,328 size 15x15
      Appearance <- "HMI_Status_G120D_Status"
   Circle "Kreis_21" at 813,353 size 15x15
      Appearance <- "HMI_Status_G120D_Status"
   Circle "Kreis_22" at 813,378 size 15x15
      Appearance <- "HMI_Status_G120D_Status"
   Circle "Kreis_23" at 813,403 size 15x15
      Appearance <- "HMI_Status_G120D_Status"
   Circle "Kreis_24" at 813,428 size 15x15
      Appearance <- "HMI_Status_G120D_Status"
   Circle "Kreis_25" at 813,453 size 15x15
      Appearance <- "HMI_Status_G120D_Status"
   Circle "Kreis_26" at 813,478 size 15x15
      Appearance <- "HMI_Status_G120D_Status"
   Circle "Kreis_27" at 813,503 size 15x15
      Appearance <- "HMI_Status_G120D_Status"
   Circle "Kreis_28" at 813,528 size 15x15
      Appearance <- "HMI_Status_G120D_Status"
   Circle "Kreis_29" at 813,553 size 15x15
      Appearance <- "HMI_Status_G120D_Status"
   Circle "Kreis_30" at 813,578 size 15x15
      Appearance <- "HMI_Status_G120D_Status"
   Circle "Kreis_31" at 813,603 size 15x15
      Appearance <- "HMI_Status_G120D_Status"
   Circle "Kreis_32" at 813,628 size 15x15
      Appearance <- "HMI_Status_G120D_Status"
   TextField "Text field_3" at 128,698 size 65x25; Text 'FAULT'
   TextField "Text field_4" at 93,743 size 100x25; Text 'WARNING'

screen "735_DIST_CONTROL_SYNCH_NOT_USED" 1280x800, template "Top_Header"
   on GenerateScreen: SetTag("SDC\_intern_Bildnummer", 735)
   Button "Schaltfläche_2" at 144,128 size 70x593; TextOff 'Text'
   Button "Schaltfläche_1" at 214,128 size 915x42; TextOff 'Text'
   IOField "EA-Feld_6" at 217,176 size 96x29; Authorization "Benutzerverwaltung"; FormatPattern 99999999
      Appearance <- "SDC\_EDIT"
      ProcessValue <- "DB_SDC_GLOBAL_SYNCH[0].HYST"
      ObjectEnable <- "SDC\_EDIT"
   TextField "Textfeld_5" at 156,179 size 35x23; Text '1'
   Button "Schaltfläche_38" at 5,388 size 127x84; TextOff 'EDIT'
      on Click: SetTag("SDC\_EDIT", 1); InvertBit("SDC\_EDIT_BIT")
      Appearance <- "SDC\_EDIT"
   TextField "Textfeld_10" at 156,213 size 35x23; Text '2'
   TextField "Textfeld_14" at 156,247 size 35x23; Text '3'
   TextField "Textfeld_15" at 156,281 size 35x23; Text '4'
   TextField "Textfeld_16" at 156,315 size 35x23; Text '5'
   TextField "Textfeld_17" at 157,349 size 35x23; Text '6'
   TextField "Textfeld_18" at 156,384 size 35x23; Text '7'
   TextField "Textfeld_19" at 156,418 size 35x23; Text '8'
   TextField "Textfeld_20" at 156,452 size 35x23; Text '9'
   TextField "Textfeld_21" at 156,486 size 35x23; Text '10'
   IOField "EA-Feld_18" at 320,176 size 64x29; Authorization "Benutzerverwaltung"; FormatPattern 99.9
      Appearance <- "SDC\_EDIT"
      ProcessValue <- "DB_SDC_GLOBAL_SYNCH[0].K"
      ObjectEnable <- "SDC\_EDIT"
   TextField "Textfeld_22" at 148,138 size 58x27; Text 'ParSet'
   TextField "Textfeld_23" at 156,520 size 35x23; Text '11'
   TextField "Textfeld_24" at 156,555 size 35x23; Text '12'
   TextField "Textfeld_25" at 156,589 size 35x23; Text '13'
   TextField "Textfeld_26" at 156,623 size 35x23; Text '14'
   TextField "Textfeld_27" at 156,657 size 35x23; Text '15'
   TextField "Textfeld_28" at 156,692 size 35x23; Text '16'
   TextField "Textfeld_34" at 221,137 size 87x27; Text 'hysterese / Hysterese / Hysteresis'
   TextField "Textfeld_35" at 315,137 size 42x27; Text 'gain / Gain'
   IOField "EA-Feld_10" at 390,176 size 64x29; Authorization "Benutzerverwaltung"; FormatPattern 99.99
      Appearance <- "SDC\_EDIT"
      ProcessValue <- "DB_SDC_GLOBAL_SYNCH[0].MAX_FAKT"
      ObjectEnable <- "SDC\_EDIT"
   IOField "EA-Feld_51" at 529,176 size 120x29; Authorization "Benutzerverwaltung"; FormatPattern 99999999
      Appearance <- "SDC\_EDIT"
      ProcessValue <- "DB_SDC_GLOBAL_SYNCH[0].SET_DIST"
      ObjectEnable <- "SDC\_EDIT"
   IOField "EA-Feld_52" at 655,176 size 120x29; Authorization "Benutzerverwaltung"; FormatPattern 99999999
      Appearance <- "SDC\_EDIT"
      ProcessValue <- "DB_SDC_GLOBAL_SYNCH[0].SYNCH_DIST"
      ObjectEnable <- "SDC\_EDIT"
   TextField "Textfeld_39" at 399,137 size 40x27; Text 'max / Max'
   IOField "EA-Feld_12" at 459,176 size 64x29; Authorization "Benutzerverwaltung"; FormatPattern 99.9
      Appearance <- "SDC\_EDIT"
      ProcessValue <- "DB_SDC_GLOBAL_SYNCH[0].MIN_FAKT"
      ObjectEnable <- "SDC\_EDIT"
   TextField "Textfeld_40" at 466,137 size 40x27; Text 'min / Min'
   TextField "Textfeld_41" at 533,137 size 93x27; Text 'setpoint / Setpoint- / / Set Point'
   TextField "Textfeld_49" at 604,137 size 155x27; Text 'start value / Start Synchron- / / Start Value'
   IOField "EA-Feld_53" at 217,210 size 96x29; Authorization "Benutzerverwaltung"; FormatPattern 99999999
      Appearance <- "SDC\_EDIT"
      ProcessValue <- "DB_SDC_GLOBAL_SYNCH[1].HYST"
      ObjectEnable <- "SDC\_EDIT"
   IOField "EA-Feld_54" at 320,210 size 64x29; Authorization "Benutzerverwaltung"; FormatPattern 99.9
      Appearance <- "SDC\_EDIT"
      ProcessValue <- "DB_SDC_GLOBAL_SYNCH[1].K"
      ObjectEnable <- "SDC\_EDIT"
   IOField "EA-Feld_55" at 390,210 size 64x29; Authorization "Benutzerverwaltung"; FormatPattern 99.99
      Appearance <- "SDC\_EDIT"
      ProcessValue <- "DB_SDC_GLOBAL_SYNCH[1].MAX_FAKT"
      ObjectEnable <- "SDC\_EDIT"
   IOField "EA-Feld_56" at 529,210 size 120x29; Authorization "Benutzerverwaltung"; FormatPattern 99999999
      Appearance <- "SDC\_EDIT"
      ProcessValue <- "DB_SDC_GLOBAL_SYNCH[1].SET_DIST"
      ObjectEnable <- "SDC\_EDIT"
   IOField "EA-Feld_57" at 655,210 size 120x29; Authorization "Benutzerverwaltung"; FormatPattern 99999999
      Appearance <- "SDC\_EDIT"
      ProcessValue <- "DB_SDC_GLOBAL_SYNCH[1].SYNCH_DIST"
      ObjectEnable <- "SDC\_EDIT"
   IOField "EA-Feld_58" at 459,210 size 64x29; Authorization "Benutzerverwaltung"; FormatPattern 99.9
      Appearance <- "SDC\_EDIT"
      ProcessValue <- "DB_SDC_GLOBAL_SYNCH[1].MIN_FAKT"
      ObjectEnable <- "SDC\_EDIT"
   IOField "EA-Feld_59" at 217,245 size 96x29; Authorization "Benutzerverwaltung"; FormatPattern 99999999
      Appearance <- "SDC\_EDIT"
      ProcessValue <- "DB_SDC_GLOBAL_SYNCH[2].HYST"
      ObjectEnable <- "SDC\_EDIT"
   IOField "EA-Feld_60" at 320,245 size 64x29; Authorization "Benutzerverwaltung"; FormatPattern 99.9
      Appearance <- "SDC\_EDIT"
      ProcessValue <- "DB_SDC_GLOBAL_SYNCH[2].K"
      ObjectEnable <- "SDC\_EDIT"
   IOField "EA-Feld_61" at 390,245 size 64x29; Authorization "Benutzerverwaltung"; FormatPattern 99.99
      Appearance <- "SDC\_EDIT"
      ProcessValue <- "DB_SDC_GLOBAL_SYNCH[2].MAX_FAKT"
      ObjectEnable <- "SDC\_EDIT"
   IOField "EA-Feld_62" at 529,245 size 120x29; Authorization "Benutzerverwaltung"; FormatPattern 99999999
      Appearance <- "SDC\_EDIT"
      ProcessValue <- "DB_SDC_GLOBAL_SYNCH[2].SET_DIST"
      ObjectEnable <- "SDC\_EDIT"
   IOField "EA-Feld_63" at 655,245 size 120x29; Authorization "Benutzerverwaltung"; FormatPattern 99999999
      Appearance <- "SDC\_EDIT"
      ProcessValue <- "DB_SDC_GLOBAL_SYNCH[2].SYNCH_DIST"
      ObjectEnable <- "SDC\_EDIT"
   IOField "EA-Feld_64" at 459,245 size 64x29; Authorization "Benutzerverwaltung"; FormatPattern 99.9
      Appearance <- "SDC\_EDIT"
      ProcessValue <- "DB_SDC_GLOBAL_SYNCH[2].MIN_FAKT"
      ObjectEnable <- "SDC\_EDIT"
   IOField "EA-Feld_65" at 217,280 size 96x29; Authorization "Benutzerverwaltung"; FormatPattern 99999999
      Appearance <- "SDC\_EDIT"
      ProcessValue <- "DB_SDC_GLOBAL_SYNCH[3].HYST"
      ObjectEnable <- "SDC\_EDIT"
   IOField "EA-Feld_66" at 320,280 size 64x29; Authorization "Benutzerverwaltung"; FormatPattern 99.9
      Appearance <- "SDC\_EDIT"
      ProcessValue <- "DB_SDC_GLOBAL_SYNCH[3].K"
      ObjectEnable <- "SDC\_EDIT"
   IOField "EA-Feld_67" at 390,280 size 64x29; Authorization "Benutzerverwaltung"; FormatPattern 99.99
      Appearance <- "SDC\_EDIT"
      ProcessValue <- "DB_SDC_GLOBAL_SYNCH[3].MAX_FAKT"
      ObjectEnable <- "SDC\_EDIT"
   IOField "EA-Feld_68" at 529,280 size 120x29; Authorization "Benutzerverwaltung"; FormatPattern 99999999
      Appearance <- "SDC\_EDIT"
      ProcessValue <- "DB_SDC_GLOBAL_SYNCH[3].SET_DIST"
      ObjectEnable <- "SDC\_EDIT"
   IOField "EA-Feld_69" at 655,280 size 120x29; Authorization "Benutzerverwaltung"; FormatPattern 99999999
      Appearance <- "SDC\_EDIT"
      ProcessValue <- "DB_SDC_GLOBAL_SYNCH[3].SYNCH_DIST"
      ObjectEnable <- "SDC\_EDIT"
   IOField "EA-Feld_70" at 459,280 size 64x29; Authorization "Benutzerverwaltung"; FormatPattern 99.9
      Appearance <- "SDC\_EDIT"
      ProcessValue <- "DB_SDC_GLOBAL_SYNCH[3].MIN_FAKT"
      ObjectEnable <- "SDC\_EDIT"
   IOField "EA-Feld_71" at 217,314 size 96x29; Authorization "Benutzerverwaltung"; FormatPattern 99999999
      Appearance <- "SDC\_EDIT"
      ProcessValue <- "DB_SDC_GLOBAL_SYNCH[4].HYST"
      ObjectEnable <- "SDC\_EDIT"
   IOField "EA-Feld_72" at 320,314 size 64x29; Authorization "Benutzerverwaltung"; FormatPattern 99.9
      Appearance <- "SDC\_EDIT"
      ProcessValue <- "DB_SDC_GLOBAL_SYNCH[4].K"
      ObjectEnable <- "SDC\_EDIT"
   IOField "EA-Feld_73" at 390,314 size 64x29; Authorization "Benutzerverwaltung"; FormatPattern 99.99
      Appearance <- "SDC\_EDIT"
      ProcessValue <- "DB_SDC_GLOBAL_SYNCH[4].MAX_FAKT"
      ObjectEnable <- "SDC\_EDIT"
   IOField "EA-Feld_74" at 529,314 size 120x29; Authorization "Benutzerverwaltung"; FormatPattern 99999999
      Appearance <- "SDC\_EDIT"
      ProcessValue <- "DB_SDC_GLOBAL_SYNCH[4].SET_DIST"
      ObjectEnable <- "SDC\_EDIT"
   IOField "EA-Feld_75" at 655,314 size 120x29; Authorization "Benutzerverwaltung"; FormatPattern 99999999
      Appearance <- "SDC\_EDIT"
      ProcessValue <- "DB_SDC_GLOBAL_SYNCH[4].SYNCH_DIST"
      ObjectEnable <- "SDC\_EDIT"
   IOField "EA-Feld_76" at 459,314 size 64x29; Authorization "Benutzerverwaltung"; FormatPattern 99.9
      Appearance <- "SDC\_EDIT"
      ProcessValue <- "DB_SDC_GLOBAL_SYNCH[4].MIN_FAKT"
      ObjectEnable <- "SDC\_EDIT"
   IOField "EA-Feld_77" at 217,349 size 96x29; Authorization "Benutzerverwaltung"; FormatPattern 99999999
      Appearance <- "SDC\_EDIT"
      ProcessValue <- "DB_SDC_GLOBAL_SYNCH[5].HYST"
      ObjectEnable <- "SDC\_EDIT"
   IOField "EA-Feld_78" at 320,349 size 64x29; Authorization "Benutzerverwaltung"; FormatPattern 99.9
      Appearance <- "SDC\_EDIT"
      ProcessValue <- "DB_SDC_GLOBAL_SYNCH[5].K"
      ObjectEnable <- "SDC\_EDIT"
   IOField "EA-Feld_79" at 390,349 size 64x29; Authorization "Benutzerverwaltung"; FormatPattern 99.99
      Appearance <- "SDC\_EDIT"
      ProcessValue <- "DB_SDC_GLOBAL_SYNCH[5].MAX_FAKT"
      ObjectEnable <- "SDC\_EDIT"
   IOField "EA-Feld_80" at 529,349 size 120x29; Authorization "Benutzerverwaltung"; FormatPattern 99999999
      Appearance <- "SDC\_EDIT"
      ProcessValue <- "DB_SDC_GLOBAL_SYNCH[5].SET_DIST"
      ObjectEnable <- "SDC\_EDIT"
   IOField "EA-Feld_81" at 655,349 size 120x29; Authorization "Benutzerverwaltung"; FormatPattern 99999999
      Appearance <- "SDC\_EDIT"
      ProcessValue <- "DB_SDC_GLOBAL_SYNCH[5].SYNCH_DIST"
      ObjectEnable <- "SDC\_EDIT"
   IOField "EA-Feld_82" at 459,349 size 64x29; Authorization "Benutzerverwaltung"; FormatPattern 99.9
      Appearance <- "SDC\_EDIT"
      ProcessValue <- "DB_SDC_GLOBAL_SYNCH[5].MIN_FAKT"
      ObjectEnable <- "SDC\_EDIT"
   IOField "EA-Feld_83" at 217,384 size 96x29; Authorization "Benutzerverwaltung"; FormatPattern 99999999
      Appearance <- "SDC\_EDIT"
      ProcessValue <- "DB_SDC_GLOBAL_SYNCH[6].HYST"
      ObjectEnable <- "SDC\_EDIT"
   IOField "EA-Feld_84" at 320,384 size 64x29; Authorization "Benutzerverwaltung"; FormatPattern 99.9
      Appearance <- "SDC\_EDIT"
      ProcessValue <- "DB_SDC_GLOBAL_SYNCH[6].K"
      ObjectEnable <- "SDC\_EDIT"
   IOField "EA-Feld_85" at 390,384 size 64x29; Authorization "Benutzerverwaltung"; FormatPattern 99.99
      Appearance <- "SDC\_EDIT"
      ProcessValue <- "DB_SDC_GLOBAL_SYNCH[6].MAX_FAKT"
      ObjectEnable <- "SDC\_EDIT"
   IOField "EA-Feld_86" at 529,384 size 120x29; Authorization "Benutzerverwaltung"; FormatPattern 99999999
      Appearance <- "SDC\_EDIT"
      ProcessValue <- "DB_SDC_GLOBAL_SYNCH[6].SET_DIST"
      ObjectEnable <- "SDC\_EDIT"
   IOField "EA-Feld_87" at 655,384 size 120x29; Authorization "Benutzerverwaltung"; FormatPattern 99999999
      Appearance <- "SDC\_EDIT"
      ProcessValue <- "DB_SDC_GLOBAL_SYNCH[6].SYNCH_DIST"
      ObjectEnable <- "SDC\_EDIT"
   IOField "EA-Feld_88" at 459,384 size 64x29; Authorization "Benutzerverwaltung"; FormatPattern 99.9
      Appearance <- "SDC\_EDIT"
      ProcessValue <- "DB_SDC_GLOBAL_SYNCH[6].MIN_FAKT"
      ObjectEnable <- "SDC\_EDIT"
   IOField "EA-Feld_89" at 217,418 size 96x29; Authorization "Benutzerverwaltung"; FormatPattern 99999999
      Appearance <- "SDC\_EDIT"
      ProcessValue <- "DB_SDC_GLOBAL_SYNCH[7].HYST"
      ObjectEnable <- "SDC\_EDIT"
   IOField "EA-Feld_90" at 320,418 size 64x29; Authorization "Benutzerverwaltung"; FormatPattern 99.9
      Appearance <- "SDC\_EDIT"
      ProcessValue <- "DB_SDC_GLOBAL_SYNCH[7].K"
      ObjectEnable <- "SDC\_EDIT"
   IOField "EA-Feld_91" at 390,418 size 64x29; Authorization "Benutzerverwaltung"; FormatPattern 99.99
      Appearance <- "SDC\_EDIT"
      ProcessValue <- "DB_SDC_GLOBAL_SYNCH[7].MAX_FAKT"
      ObjectEnable <- "SDC\_EDIT"
   IOField "EA-Feld_92" at 529,418 size 120x29; Authorization "Benutzerverwaltung"; FormatPattern 99999999
      Appearance <- "SDC\_EDIT"
      ProcessValue <- "DB_SDC_GLOBAL_SYNCH[7].SET_DIST"
      ObjectEnable <- "SDC\_EDIT"
   IOField "EA-Feld_93" at 655,418 size 120x29; Authorization "Benutzerverwaltung"; FormatPattern 99999999
      Appearance <- "SDC\_EDIT"
      ProcessValue <- "DB_SDC_GLOBAL_SYNCH[7].SYNCH_DIST"
      ObjectEnable <- "SDC\_EDIT"
   IOField "EA-Feld_94" at 459,418 size 64x29; Authorization "Benutzerverwaltung"; FormatPattern 99.9